
   //Update XCUT status
   "FB_BPSEthLink_ServerA_V1_00_IDB".IN_rgtStatusXCuts[0].dActualCarriagePos_cmm := "FB_CrossCuts_1_V1_00_IDB".tHMR.dCarriagePosition_cmm;
   "FB_BPSEthLink_ServerA_V1_00_IDB".IN_rgtStatusXCuts[0].dDistanceFromSnaproll_cmm := "FB_CrossCuts_1_V1_00_IDB".tHMR.dDistanceFromSnaproll_cmm;
   "FB_BPSEthLink_ServerA_V1_00_IDB".IN_rgtStatusXCuts[0].dStatus := "FB_CrossCuts_1_V1_00_IDB".tHMR.dStatus;
   "FB_BPSEthLink_ServerA_V1_00_IDB".IN_rgtStatusXCuts[0].dXCutActualStatus := "FB_CrossCuts_1_V1_00_IDB".tHMR.dXCutActualStatus;
   IF "FB_CrossCuts_1_V1_00_IDB".tHMR.dXCutActualStatus = 1 THEN
       "FB_BPSEthLink_ServerA_V1_00_IDB".IN_rgtStatusXCuts[0].dStatus := 7;
   END_IF;

   "FB_BPSEthLink_ServerA_V1_00_IDB".IN_rgtStatusXCuts[1].dActualCarriagePos_cmm := "FB_CrossCuts_2_V1_00_IDB".tHMR.dCarriagePosition_cmm;
   "FB_BPSEthLink_ServerA_V1_00_IDB".IN_rgtStatusXCuts[1].dDistanceFromSnaproll_cmm := "FB_CrossCuts_2_V1_00_IDB".tHMR.dDistanceFromSnaproll_cmm;
   "FB_BPSEthLink_ServerA_V1_00_IDB".IN_rgtStatusXCuts[1].dStatus := "FB_CrossCuts_2_V1_00_IDB".tHMR.dStatus;
   "FB_BPSEthLink_ServerA_V1_00_IDB".IN_rgtStatusXCuts[1].dXCutActualStatus := "FB_CrossCuts_2_V1_00_IDB".tHMR.dXCutActualStatus;

   IF "FB_CrossCuts_2_V1_00_IDB".tHMR.dXCutActualStatus = 1 THEN
       "FB_BPSEthLink_ServerA_V1_00_IDB".IN_rgtStatusXCuts[1].dStatus := 7;
   END_IF;

   //Update YCUT status 
   "FB_BPSEthLink_ServerA_V1_00_IDB".IN_rgtStatusYCuts[0].dBridgeStatus := "FB_YCuts1_V1_00_IDB".OUT_tBridgeStatus.dBridgeStatus;
   "FB_BPSEthLink_ServerA_V1_00_IDB".IN_rgtStatusYCuts[0].dDistanceSnapRoll_cmm := "FB_YCuts1_V1_00_IDB".tHMR.dDistanceFromSnaproll_cmm;
   "FB_BPSEthLink_ServerA_V1_00_IDB".IN_rgtStatusYCuts[0].rgdPosition_cmm := "FB_YCuts1_V1_00_IDB".OUT_tBridgeStatus.rgdPosition_cmm;
   "FB_BPSEthLink_ServerA_V1_00_IDB".IN_rgtStatusYCuts[0].rgxFireON := "FB_YCuts1_V1_00_IDB".OUT_tBridgeStatus.rgxFireON;
   "FB_BPSEthLink_ServerA_V1_00_IDB".IN_rgtStatusYCuts[0].rgxHeadProdOn := "FB_YCuts1_V1_00_IDB".OUT_tBridgeStatus.rgxHeadProdOn;

   "FB_BPSEthLink_ServerA_V1_00_IDB".IN_rgtStatusYCuts[1].dBridgeStatus := "FB_YCuts2_V1_00_IDB".OUT_tBridgeStatus.dBridgeStatus;
   "FB_BPSEthLink_ServerA_V1_00_IDB".IN_rgtStatusYCuts[1].dDistanceSnapRoll_cmm := "FB_YCuts2_V1_00_IDB".tHMR.dDistanceFromSnaproll_cmm;
   "FB_BPSEthLink_ServerA_V1_00_IDB".IN_rgtStatusYCuts[1].rgdPosition_cmm := "FB_YCuts2_V1_00_IDB".OUT_tBridgeStatus.rgdPosition_cmm;
   "FB_BPSEthLink_ServerA_V1_00_IDB".IN_rgtStatusYCuts[1].rgxFireON := "FB_YCuts2_V1_00_IDB".OUT_tBridgeStatus.rgxFireON;
   "FB_BPSEthLink_ServerA_V1_00_IDB".IN_rgtStatusYCuts[1].rgxHeadProdOn := "FB_YCuts2_V1_00_IDB".OUT_tBridgeStatus.rgxHeadProdOn;

   //Update general status
   IF (("Z201".ST_xThisPlcActive) AND ("Z201".ST_xPLC1)) THEN
       "FB_BPSEthLink_ServerA_V1_00_IDB".IN_tStatusGeneral.dActivePLC := 1;
   ELSE
       "FB_BPSEthLink_ServerA_V1_00_IDB".IN_tStatusGeneral.dActivePLC := 2;
   END_IF;

   "FB_BPSEthLink_ServerA_V1_00_IDB".IN_tStatusGeneral.dAutoRibSelection := "FB_OptManager_V1_00_IDB".tHMW.dSelectWanderDataSource;
   "FB_BPSEthLink_ServerA_V1_00_IDB".IN_tStatusGeneral.dExtOptSelected := "FB_OptManager_V1_00_IDB".tHMR.dSelOptimizer;
   "FB_BPSEthLink_ServerA_V1_00_IDB".IN_tStatusGeneral.dOptimizerMode := 2;

   IF "FB_OptEthLink_V1_00_IDB".tALM.tS.xCh1NotCon AND "FB_OptEthLink_V1_00_IDB".tALM.tS.xCh2NotCon THEN 
       "FB_BPSEthLink_ServerA_V1_00_IDB".IN_tStatusGeneral.dOptStatus := 1;
   ELSIF "FB_OptEthLink_V1_00_IDB".tALM.tS.xCh1NotCon OR "FB_OptEthLink_V1_00_IDB".tALM.tS.xCh2NotCon THEN
       "FB_BPSEthLink_ServerA_V1_00_IDB".IN_tStatusGeneral.dOptStatus := 7;
   ELSE
       "FB_BPSEthLink_ServerA_V1_00_IDB".IN_tStatusGeneral.dOptStatus := 3;
   END_IF;

   IF "FB_OptManager_V1_00_IDB".tHMW.dSelectWanderDataSource > 0 THEN
       "FB_BPSEthLink_ServerA_V1_00_IDB".IN_tStatusGeneral.dRibbonModality := 1;
   ELSE
       "FB_BPSEthLink_ServerA_V1_00_IDB".IN_tStatusGeneral.dRibbonModality := 4;
   END_IF;

   "FB_BPSEthLink_ServerA_V1_00_IDB".IN_tStatusGeneral.dScanStatus := "FB_ISRA5D_IDB".tHMR.dInspectionStatus;

   IF "FB_OptManager_V1_00_IDB".tHMW.dSelectWanderMode = 0 THEN
       "FB_BPSEthLink_ServerA_V1_00_IDB".IN_tStatusGeneral.dTypeWanderSel := 2;
   ELSE
       "FB_BPSEthLink_ServerA_V1_00_IDB".IN_tStatusGeneral.dTypeWanderSel := 1;
   END_IF;

   "FB_BPSEthLink_ServerA_V1_00_IDB".IN_tStatusGeneral.dYC1WandRec_cmm := "FB_YCuts1_V1_00_IDB".AUX_dActualRecoverWander_cmm;
   "FB_BPSEthLink_ServerA_V1_00_IDB".IN_tStatusGeneral.dYC2WandRec_cmm := "FB_YCuts2_V1_00_IDB".AUX_dActualRecoverWander_cmm;
   "FB_BPSEthLink_ServerA_V1_00_IDB".IN_tStatusGeneral.dWanderRecoveryThr_cmm := "FB_OptManager_V1_00_IDB".tHMW.dWanderRecThr_cmm;

   "FB_BPSEthLink_ServerA_V1_00_IDB".IN_tStatusGeneral.dScanGrossWidth_cmm := "FB_ISRA5D_IDB".tHMR.dCurrentGrossWidth_cmm;
   "FB_BPSEthLink_ServerA_V1_00_IDB".IN_tStatusGeneral.dScanNetWidth_cmm := "FB_ISRA5D_IDB".tHMR.dCurrentNetWidth_cmm;
   "FB_BPSEthLink_ServerA_V1_00_IDB".IN_tStatusGeneral.dScanGrossWander_cmm := "FB_ISRA5D_IDB".tHMR.dCurrentGrossWander_cmm;
   "FB_BPSEthLink_ServerA_V1_00_IDB".IN_tStatusGeneral.dScanNetWander_cmm := "FB_ISRA5D_IDB".tHMR.dCurrentNetWander_cmm;

   "FB_BPSEthLink_ServerA_V1_00_IDB".IN_tStatusGeneral.dCameraGrossWidth_cmm := 0;
   "FB_BPSEthLink_ServerA_V1_00_IDB".IN_tStatusGeneral.dCameraNetWidth_cmm := 0;
   "FB_BPSEthLink_ServerA_V1_00_IDB".IN_tStatusGeneral.dCameraGrossWander_cmm := 0;
   "FB_BPSEthLink_ServerA_V1_00_IDB".IN_tStatusGeneral.dCameraNetWander_cmm := 0;



   //BPS Connection B

   "FB_BPSEthLink_ServerB_V1_00_IDB".IN_tRemoteAddress.ADDR[1] := "IPV4_BPS_SERVERB_IP1";
   "FB_BPSEthLink_ServerB_V1_00_IDB".IN_tRemoteAddress.ADDR[2] := "IPV4_BPS_SERVERB_IP2";
   "FB_BPSEthLink_ServerB_V1_00_IDB".IN_tRemoteAddress.ADDR[3] := "IPV4_BPS_SERVERB_IP3";
   "FB_BPSEthLink_ServerB_V1_00_IDB".IN_tRemoteAddress.ADDR[4] := "IPV4_BPS_SERVERB_IP4";

   "FB_BPSEthLink_ServerB_V1_00_IDB".IN_tStatusEncoder.dActualBTC_cmm := "DB_Encoder".dActualEncoderCounter_cmm;
   "FB_BPSEthLink_ServerB_V1_00_IDB".IN_tStatusEncoder.dTrackSpeed_mm_min := "DB_Encoder".dActSpeedValue_mm_min;

   //Update XCUT status
   "FB_BPSEthLink_ServerB_V1_00_IDB".IN_rgtStatusXCuts[0].dActualCarriagePos_cmm := "FB_CrossCuts_1_V1_00_IDB".tHMR.dCarriagePosition_cmm;
   "FB_BPSEthLink_ServerB_V1_00_IDB".IN_rgtStatusXCuts[0].dDistanceFromSnaproll_cmm := "FB_CrossCuts_1_V1_00_IDB".tHMR.dDistanceFromSnaproll_cmm;
   "FB_BPSEthLink_ServerB_V1_00_IDB".IN_rgtStatusXCuts[0].dStatus := "FB_CrossCuts_1_V1_00_IDB".tHMR.dStatus;
   "FB_BPSEthLink_ServerB_V1_00_IDB".IN_rgtStatusXCuts[0].dXCutActualStatus := "FB_CrossCuts_1_V1_00_IDB".tHMR.dXCutActualStatus;

   IF "FB_CrossCuts_1_V1_00_IDB".tHMR.dXCutActualStatus = 1 THEN
       "FB_BPSEthLink_ServerB_V1_00_IDB".IN_rgtStatusXCuts[0].dStatus := 7;
   END_IF;

   "FB_BPSEthLink_ServerB_V1_00_IDB".IN_rgtStatusXCuts[1].dActualCarriagePos_cmm := "FB_CrossCuts_2_V1_00_IDB".tHMR.dCarriagePosition_cmm;
   "FB_BPSEthLink_ServerB_V1_00_IDB".IN_rgtStatusXCuts[1].dDistanceFromSnaproll_cmm := "FB_CrossCuts_2_V1_00_IDB".tHMR.dDistanceFromSnaproll_cmm;
   "FB_BPSEthLink_ServerB_V1_00_IDB".IN_rgtStatusXCuts[1].dStatus := "FB_CrossCuts_2_V1_00_IDB".tHMR.dStatus;
   "FB_BPSEthLink_ServerB_V1_00_IDB".IN_rgtStatusXCuts[1].dXCutActualStatus := "FB_CrossCuts_2_V1_00_IDB".tHMR.dXCutActualStatus;

   IF "FB_CrossCuts_2_V1_00_IDB".tHMR.dXCutActualStatus = 1 THEN
       "FB_BPSEthLink_ServerB_V1_00_IDB".IN_rgtStatusXCuts[1].dStatus := 7;
   END_IF;

   //Update YCUT status 
   "FB_BPSEthLink_ServerB_V1_00_IDB".IN_rgtStatusYCuts[0].dBridgeStatus := "FB_YCuts1_V1_00_IDB".OUT_tBridgeStatus.dBridgeStatus;
   "FB_BPSEthLink_ServerB_V1_00_IDB".IN_rgtStatusYCuts[0].dDistanceSnapRoll_cmm := "FB_YCuts1_V1_00_IDB".tHMR.dDistanceFromSnaproll_cmm;
   "FB_BPSEthLink_ServerB_V1_00_IDB".IN_rgtStatusYCuts[0].rgdPosition_cmm := "FB_YCuts1_V1_00_IDB".OUT_tBridgeStatus.rgdPosition_cmm;
   "FB_BPSEthLink_ServerB_V1_00_IDB".IN_rgtStatusYCuts[0].rgxFireON := "FB_YCuts1_V1_00_IDB".OUT_tBridgeStatus.rgxFireON;
   "FB_BPSEthLink_ServerB_V1_00_IDB".IN_rgtStatusYCuts[0].rgxHeadProdOn := "FB_YCuts1_V1_00_IDB".OUT_tBridgeStatus.rgxHeadProdOn;

   "FB_BPSEthLink_ServerB_V1_00_IDB".IN_rgtStatusYCuts[1].dBridgeStatus := "FB_YCuts2_V1_00_IDB".OUT_tBridgeStatus.dBridgeStatus;
   "FB_BPSEthLink_ServerB_V1_00_IDB".IN_rgtStatusYCuts[1].dDistanceSnapRoll_cmm := "FB_YCuts2_V1_00_IDB".tHMR.dDistanceFromSnaproll_cmm;
   "FB_BPSEthLink_ServerB_V1_00_IDB".IN_rgtStatusYCuts[1].rgdPosition_cmm := "FB_YCuts2_V1_00_IDB".OUT_tBridgeStatus.rgdPosition_cmm;
   "FB_BPSEthLink_ServerB_V1_00_IDB".IN_rgtStatusYCuts[1].rgxFireON := "FB_YCuts2_V1_00_IDB".OUT_tBridgeStatus.rgxFireON;
   "FB_BPSEthLink_ServerB_V1_00_IDB".IN_rgtStatusYCuts[1].rgxHeadProdOn := "FB_YCuts2_V1_00_IDB".OUT_tBridgeStatus.rgxHeadProdOn;

   //Update general status
   IF (("Z201".ST_xThisPlcActive) AND ("Z201".ST_xPLC1)) THEN
       "FB_BPSEthLink_ServerB_V1_00_IDB".IN_tStatusGeneral.dActivePLC := 1;
   ELSE
       "FB_BPSEthLink_ServerB_V1_00_IDB".IN_tStatusGeneral.dActivePLC := 2;
   END_IF;

   "FB_BPSEthLink_ServerB_V1_00_IDB".IN_tStatusGeneral.dAutoRibSelection := "FB_OptManager_V1_00_IDB".tHMW.dSelectWanderDataSource;
   "FB_BPSEthLink_ServerB_V1_00_IDB".IN_tStatusGeneral.dExtOptSelected := "FB_OptManager_V1_00_IDB".tHMR.dSelOptimizer;
   "FB_BPSEthLink_ServerB_V1_00_IDB".IN_tStatusGeneral.dOptimizerMode := 2;

   IF "FB_OptEthLink_V1_00_IDB".tALM.tS.xCh1NotCon AND "FB_OptEthLink_V1_00_IDB".tALM.tS.xCh2NotCon THEN 
       "FB_BPSEthLink_ServerB_V1_00_IDB".IN_tStatusGeneral.dOptStatus := 1;
   ELSIF "FB_OptEthLink_V1_00_IDB".tALM.tS.xCh1NotCon OR "FB_OptEthLink_V1_00_IDB".tALM.tS.xCh2NotCon THEN
       "FB_BPSEthLink_ServerB_V1_00_IDB".IN_tStatusGeneral.dOptStatus := 7;
   ELSE
       "FB_BPSEthLink_ServerB_V1_00_IDB".IN_tStatusGeneral.dOptStatus := 3;
   END_IF;

   IF "FB_OptManager_V1_00_IDB".tHMW.dSelectWanderDataSource > 0 THEN
       "FB_BPSEthLink_ServerB_V1_00_IDB".IN_tStatusGeneral.dRibbonModality := 1;
   ELSE
       "FB_BPSEthLink_ServerB_V1_00_IDB".IN_tStatusGeneral.dRibbonModality := 4;
   END_IF;

   "FB_BPSEthLink_ServerB_V1_00_IDB".IN_tStatusGeneral.dScanStatus := "FB_ISRA5D_IDB".tHMR.dInspectionStatus;

   IF "FB_OptManager_V1_00_IDB".tHMW.dSelectWanderMode = 0 THEN
       "FB_BPSEthLink_ServerB_V1_00_IDB".IN_tStatusGeneral.dTypeWanderSel := 2;
   ELSE
       "FB_BPSEthLink_ServerB_V1_00_IDB".IN_tStatusGeneral.dTypeWanderSel := 1;
   END_IF;

   "FB_BPSEthLink_ServerB_V1_00_IDB".IN_tStatusGeneral.dYC1WandRec_cmm := "FB_YCuts1_V1_00_IDB".AUX_dActualRecoverWander_cmm;
   "FB_BPSEthLink_ServerB_V1_00_IDB".IN_tStatusGeneral.dYC2WandRec_cmm := "FB_YCuts2_V1_00_IDB".AUX_dActualRecoverWander_cmm;
   "FB_BPSEthLink_ServerB_V1_00_IDB".IN_tStatusGeneral.dWanderRecoveryThr_cmm := "FB_OptManager_V1_00_IDB".tHMW.dWanderRecThr_cmm;

   "FB_BPSEthLink_ServerB_V1_00_IDB".IN_tStatusGeneral.dScanGrossWidth_cmm := "FB_ISRA5D_IDB".tHMR.dCurrentGrossWidth_cmm;
   "FB_BPSEthLink_ServerB_V1_00_IDB".IN_tStatusGeneral.dScanNetWidth_cmm := "FB_ISRA5D_IDB".tHMR.dCurrentNetWidth_cmm;
   "FB_BPSEthLink_ServerB_V1_00_IDB".IN_tStatusGeneral.dScanGrossWander_cmm := "FB_ISRA5D_IDB".tHMR.dCurrentGrossWander_cmm;
   "FB_BPSEthLink_ServerB_V1_00_IDB".IN_tStatusGeneral.dScanNetWander_cmm := "FB_ISRA5D_IDB".tHMR.dCurrentNetWander_cmm;

   "FB_BPSEthLink_ServerB_V1_00_IDB".IN_tStatusGeneral.dCameraGrossWidth_cmm := 0;
   "FB_BPSEthLink_ServerB_V1_00_IDB".IN_tStatusGeneral.dCameraNetWidth_cmm := 0;
   "FB_BPSEthLink_ServerB_V1_00_IDB".IN_tStatusGeneral.dCameraGrossWander_cmm := 0;
   "FB_BPSEthLink_ServerB_V1_00_IDB".IN_tStatusGeneral.dCameraNetWander_cmm := 0;
END_REGION

REGION Network 4: BPS A Connection data
   RUNG wire#powerrail
      "FB_BPSEthLink_ServerA_V1_00_IDB"(IN_xBPSServerA := TRUE, IN_xCycleON :=, IN_xCycleONDel := "Z201".ST_xCycleONDelayed, IN_xGeneralReset := "Z201".ST_xMachineReset, IN_xResetAlarms := "Z201".tmOFF_ResetAlarm.OUT_xDone, IN_xFaultsEnabled := "Z201".ST_xFaultsEnabled, IN_xThisPLCActive := "Z201".ST_xThisPlcActive, IN_dLineSpeed_mm_min := "FB_CommunicationZ300_V1.00_DB".IN_tIDeviceDataIN.Z300.dLineSpeed_mm_min, IN_tStatusGeneral :=, IN_tStatusEncoder :=, IN_tStatusDigitizer_1 :=, IN_tStatusDigitizer_2 :=, IN_rgtStatusXCuts :=, IN_rgtStatusYCuts :=, IN_rgtStatusMarkers :=, IN_tInterfaceID := "Local~PROFINET_MCC1200", IN_tID := "CONNUOC_BPS_SERVERA", IN_tRemoteAddress :=, IN_uiRemotePort := "UINT_BPS_SERVERA_PORT", INO_tCaps := "DB_Plates", INO_tInitialize := "GP_OB_Initialize_Main_IDB", INO_tDefects := "DB_Defects".THIS, INO_tMessages := "RP_Message".tTankMessageForReport, INO_tAddMessageFromOpt := "RP_Message".MexFromOptimizer.tAddMessageFromOptTaskMain, INO_tRibbon := "DB_RibbonData", INO_xMessageAnomaly := "RP_Message".tALM.tS.xMessageAnomaly)
   END_RUNG
   // the same network as SCL:
   "FB_BPSEthLink_ServerA_V1_00_IDB"(IN_xBPSServerA := TRUE,   // "FB_BPSEthLink_V1.00"
                           IN_xCycleONDel := "Z201".ST_xCycleONDelayed,
                           IN_xGeneralReset := "Z201".ST_xMachineReset,
                           IN_xResetAlarms := "Z201".tmOFF_ResetAlarm.OUT_xDone,
                           IN_xFaultsEnabled := "Z201".ST_xFaultsEnabled,
                           IN_xThisPLCActive := "Z201".ST_xThisPlcActive,
                           IN_dLineSpeed_mm_min := "FB_CommunicationZ300_V1.00_DB".IN_tIDeviceDataIN.Z300.dLineSpeed_mm_min,
                           IN_tInterfaceID := "Local~PROFINET_MCC1200",
                           IN_tID := "CONNUOC_BPS_SERVERA",
                           IN_uiRemotePort := "UINT_BPS_SERVERA_PORT",
                           INO_tCaps := "DB_Plates",
                           INO_tInitialize := "GP_OB_Initialize_Main_IDB",
                           INO_tDefects := "DB_Defects".THIS,
                           INO_tMessages := "RP_Message".tTankMessageForReport,
                           INO_tAddMessageFromOpt := "RP_Message".MexFromOptimizer.tAddMessageFromOptTaskMain,
                           INO_tRibbon := "DB_RibbonData",
                           INO_xMessageAnomaly := "RP_Message".tALM.tS.xMessageAnomaly);
END_REGION

REGION Network 5: BPS B Connection data
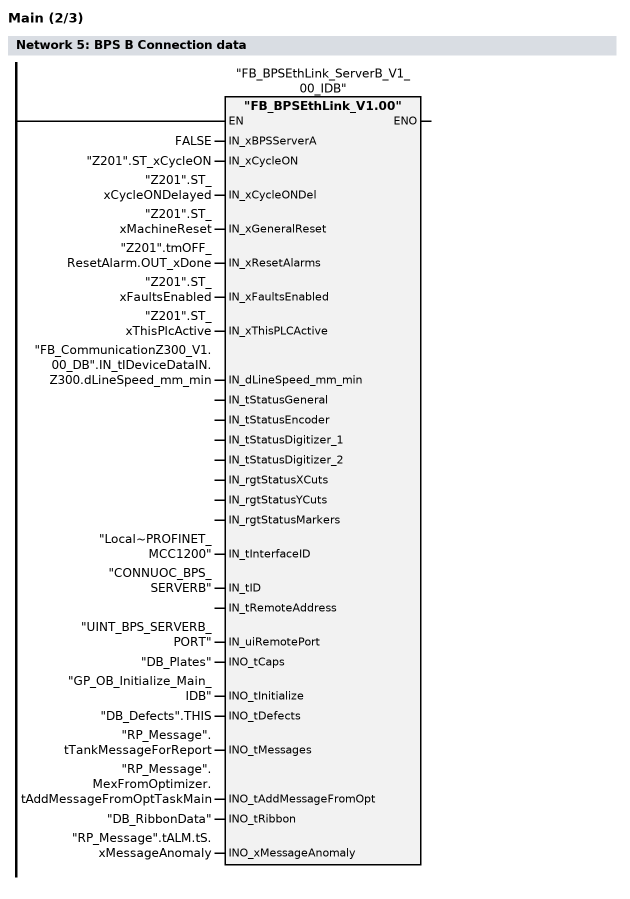
   RUNG wire#powerrail
      "FB_BPSEthLink_ServerB_V1_00_IDB"(IN_xBPSServerA := FALSE, IN_xCycleON := "Z201".ST_xCycleON, IN_xCycleONDel := "Z201".ST_xCycleONDelayed, IN_xGeneralReset := "Z201".ST_xMachineReset, IN_xResetAlarms := "Z201".tmOFF_ResetAlarm.OUT_xDone, IN_xFaultsEnabled := "Z201".ST_xFaultsEnabled, IN_xThisPLCActive := "Z201".ST_xThisPlcActive, IN_dLineSpeed_mm_min := "FB_CommunicationZ300_V1.00_DB".IN_tIDeviceDataIN.Z300.dLineSpeed_mm_min, IN_tStatusGeneral :=, IN_tStatusEncoder :=, IN_tStatusDigitizer_1 :=, IN_tStatusDigitizer_2 :=, IN_rgtStatusXCuts :=, IN_rgtStatusYCuts :=, IN_rgtStatusMarkers :=, IN_tInterfaceID := "Local~PROFINET_MCC1200", IN_tID := "CONNUOC_BPS_SERVERB", IN_tRemoteAddress :=, IN_uiRemotePort := "UINT_BPS_SERVERB_PORT", INO_tCaps := "DB_Plates", INO_tInitialize := "GP_OB_Initialize_Main_IDB", INO_tDefects := "DB_Defects".THIS, INO_tMessages := "RP_Message".tTankMessageForReport, INO_tAddMessageFromOpt := "RP_Message".MexFromOptimizer.tAddMessageFromOptTaskMain, INO_tRibbon := "DB_RibbonData", INO_xMessageAnomaly := "RP_Message".tALM.tS.xMessageAnomaly)
   END_RUNG
   // the same network as SCL:
   "FB_BPSEthLink_ServerB_V1_00_IDB"(IN_xBPSServerA := FALSE,   // "FB_BPSEthLink_V1.00"
                           IN_xCycleON := "Z201".ST_xCycleON,
                           IN_xCycleONDel := "Z201".ST_xCycleONDelayed,
                           IN_xGeneralReset := "Z201".ST_xMachineReset,
                           IN_xResetAlarms := "Z201".tmOFF_ResetAlarm.OUT_xDone,
                           IN_xFaultsEnabled := "Z201".ST_xFaultsEnabled,
                           IN_xThisPLCActive := "Z201".ST_xThisPlcActive,
                           IN_dLineSpeed_mm_min := "FB_CommunicationZ300_V1.00_DB".IN_tIDeviceDataIN.Z300.dLineSpeed_mm_min,
                           IN_tInterfaceID := "Local~PROFINET_MCC1200",
                           IN_tID := "CONNUOC_BPS_SERVERB",
                           IN_uiRemotePort := "UINT_BPS_SERVERB_PORT",
                           INO_tCaps := "DB_Plates",
                           INO_tInitialize := "GP_OB_Initialize_Main_IDB",
                           INO_tDefects := "DB_Defects".THIS,
                           INO_tMessages := "RP_Message".tTankMessageForReport,
                           INO_tAddMessageFromOpt := "RP_Message".MexFromOptimizer.tAddMessageFromOptTaskMain,
                           INO_tRibbon := "DB_RibbonData",
                           INO_xMessageAnomaly := "RP_Message".tALM.tS.xMessageAnomaly);
END_REGION

REGION Network 6 (SCL): Optimizer connection data
   //Update YCUT status 
   "FB_OptEthLink_V1_00_IDB".IN_rgtStatusYCuts[0].dBridgeStatus := "FB_YCuts1_V1_00_IDB".OUT_tBridgeStatus.dBridgeStatus;
   "FB_OptEthLink_V1_00_IDB".IN_rgtStatusYCuts[0].dDistanceSnapRoll_cmm := "FB_YCuts1_V1_00_IDB".tHMR.dDistanceFromSnaproll_cmm;
   "FB_OptEthLink_V1_00_IDB".IN_rgtStatusYCuts[0].rgdPosition_cmm := "FB_YCuts1_V1_00_IDB".OUT_tBridgeStatus.rgdPosition_cmm;
   "FB_OptEthLink_V1_00_IDB".IN_rgtStatusYCuts[0].rgxFireON := "FB_YCuts1_V1_00_IDB".OUT_tBridgeStatus.rgxFireON;
   "FB_OptEthLink_V1_00_IDB".IN_rgtStatusYCuts[0].rgxHeadProdOn := "FB_YCuts1_V1_00_IDB".OUT_tBridgeStatus.rgxHeadProdOn;


   "FB_OptEthLink_V1_00_IDB".IN_rgtStatusYCuts[1].dBridgeStatus := "FB_YCuts2_V1_00_IDB".OUT_tBridgeStatus.dBridgeStatus;
   "FB_OptEthLink_V1_00_IDB".IN_rgtStatusYCuts[1].dDistanceSnapRoll_cmm := "FB_YCuts2_V1_00_IDB".tHMR.dDistanceFromSnaproll_cmm;
   "FB_OptEthLink_V1_00_IDB".IN_rgtStatusYCuts[1].rgdPosition_cmm := "FB_YCuts2_V1_00_IDB".OUT_tBridgeStatus.rgdPosition_cmm;
   "FB_OptEthLink_V1_00_IDB".IN_rgtStatusYCuts[1].rgxFireON := "FB_YCuts2_V1_00_IDB".OUT_tBridgeStatus.rgxFireON;
   "FB_OptEthLink_V1_00_IDB".IN_rgtStatusYCuts[1].rgxHeadProdOn := "FB_YCuts2_V1_00_IDB".OUT_tBridgeStatus.rgxHeadProdOn;
   "FB_OptEthLink_V1_00_IDB".IN_rgtStatusXCuts[0].dActualCarriagePos_cmm := "FB_CrossCuts_1_V1_00_IDB".tHMR.dCarriagePosition_cmm;
   "FB_OptEthLink_V1_00_IDB".IN_rgtStatusXCuts[0].dDistanceFromSnaproll_cmm := "FB_CrossCuts_1_V1_00_IDB".tHMR.dDistanceFromSnaproll_cmm;
   "FB_OptEthLink_V1_00_IDB".IN_rgtStatusXCuts[0].dStatus := "FB_CrossCuts_1_V1_00_IDB".tHMR.dStatus;
   "FB_OptEthLink_V1_00_IDB".IN_rgtStatusXCuts[0].dXCutActualStatus := "FB_CrossCuts_1_V1_00_IDB".tHMR.dXCutActualStatus;
   "FB_OptEthLink_V1_00_IDB".IN_rgtStatusXCuts[0].dCutTime_ms := "FB_CrossCuts_1_V1_00_IDB".AUX_dCutTime100Per_ms;

   "FB_OptEthLink_V1_00_IDB".IN_rgtStatusXCuts[1].dActualCarriagePos_cmm := "FB_CrossCuts_2_V1_00_IDB".tHMR.dCarriagePosition_cmm;
   "FB_OptEthLink_V1_00_IDB".IN_rgtStatusXCuts[1].dDistanceFromSnaproll_cmm := "FB_CrossCuts_2_V1_00_IDB".tHMR.dDistanceFromSnaproll_cmm;
   "FB_OptEthLink_V1_00_IDB".IN_rgtStatusXCuts[1].dStatus := "FB_CrossCuts_2_V1_00_IDB".tHMR.dStatus;
   "FB_OptEthLink_V1_00_IDB".IN_rgtStatusXCuts[1].dXCutActualStatus := "FB_CrossCuts_2_V1_00_IDB".tHMR.dXCutActualStatus;
   "FB_OptEthLink_V1_00_IDB".IN_rgtStatusXCuts[1].dCutTime_ms := "FB_CrossCuts_2_V1_00_IDB".AUX_dCutTime100Per_ms;

   "FB_OptEthLink_V1_00_IDB".IN_rgtStatusXCuts[2].dActualCarriagePos_cmm := 0;
   "FB_OptEthLink_V1_00_IDB".IN_rgtStatusXCuts[2].dDistanceFromSnaproll_cmm := 0;
   "FB_OptEthLink_V1_00_IDB".IN_rgtStatusXCuts[2].dStatus := 1;
   "FB_OptEthLink_V1_00_IDB".IN_rgtStatusXCuts[2].dXCutActualStatus := 1;
   "FB_OptEthLink_V1_00_IDB".IN_rgtStatusXCuts[2].dCutTime_ms := 0;

   "FB_OptEthLink_V1_00_IDB".IN_rgtStatusXCuts[3].dActualCarriagePos_cmm := 0;
   "FB_OptEthLink_V1_00_IDB".IN_rgtStatusXCuts[3].dDistanceFromSnaproll_cmm := 0;
   "FB_OptEthLink_V1_00_IDB".IN_rgtStatusXCuts[3].dStatus :=1;
   "FB_OptEthLink_V1_00_IDB".IN_rgtStatusXCuts[3].dXCutActualStatus := 1;
   "FB_OptEthLink_V1_00_IDB".IN_rgtStatusXCuts[3].dCutTime_ms := 0;

   "FB_OptEthLink_V1_00_IDB".IN_rgtStatusMarker[3].dBridgeProdModeActual := 0;
   "FB_OptEthLink_V1_00_IDB".IN_rgtStatusMarker[3].dDistanceFromCenterLine_cmm := 0;
   "FB_OptEthLink_V1_00_IDB".IN_rgtStatusMarker[3].dDistanceFromSnaproll_cmm := 0;
   "FB_OptEthLink_V1_00_IDB".IN_rgtStatusMarker[3].dHeadPosition_cmm := 0;
   "FB_OptEthLink_V1_00_IDB".IN_rgtStatusMarker[3].dSpraySpace_cmm := 0;

   "FB_OptEthLink_V1_00_IDB".IN_rgtStatusMarker[4].dBridgeProdModeActual := 0;
   "FB_OptEthLink_V1_00_IDB".IN_rgtStatusMarker[4].dDistanceFromCenterLine_cmm := 0;
   "FB_OptEthLink_V1_00_IDB".IN_rgtStatusMarker[4].dDistanceFromSnaproll_cmm := 0;
   "FB_OptEthLink_V1_00_IDB".IN_rgtStatusMarker[4].dHeadPosition_cmm := 0;
   "FB_OptEthLink_V1_00_IDB".IN_rgtStatusMarker[4].dSpraySpace_cmm := 0;
END_REGION

REGION Network 7: Optimizer connection
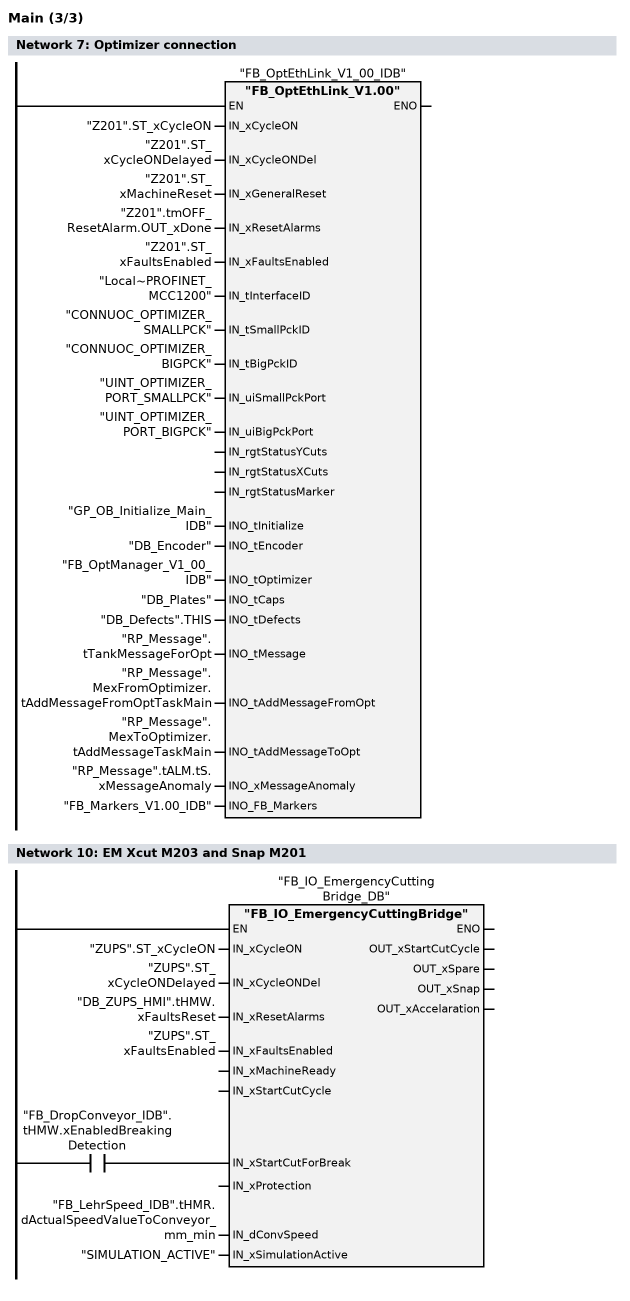
   RUNG wire#powerrail
      "FB_OptEthLink_V1_00_IDB"(IN_xCycleON := "Z201".ST_xCycleON, IN_xCycleONDel := "Z201".ST_xCycleONDelayed, IN_xGeneralReset := "Z201".ST_xMachineReset, IN_xResetAlarms := "Z201".tmOFF_ResetAlarm.OUT_xDone, IN_xFaultsEnabled := "Z201".ST_xFaultsEnabled, IN_tInterfaceID := "Local~PROFINET_MCC1200", IN_tSmallPckID := "CONNUOC_OPTIMIZER_SMALLPCK", IN_tBigPckID := "CONNUOC_OPTIMIZER_BIGPCK", IN_uiSmallPckPort := "UINT_OPTIMIZER_PORT_SMALLPCK", IN_uiBigPckPort := "UINT_OPTIMIZER_PORT_BIGPCK", IN_rgtStatusYCuts :=, IN_rgtStatusXCuts :=, IN_rgtStatusMarker :=, INO_tInitialize := "GP_OB_Initialize_Main_IDB", INO_tEncoder := "DB_Encoder", INO_tOptimizer := "FB_OptManager_V1_00_IDB", INO_tCaps := "DB_Plates", INO_tDefects := "DB_Defects".THIS, INO_tMessage := "RP_Message".tTankMessageForOpt, INO_tAddMessageFromOpt := "RP_Message".MexFromOptimizer.tAddMessageFromOptTaskMain, INO_tAddMessageToOpt := "RP_Message".MexToOptimizer.tAddMessageTaskMain, INO_xMessageAnomaly := "RP_Message".tALM.tS.xMessageAnomaly, INO_FB_Markers := "FB_Markers_V1.00_IDB")
   END_RUNG
   // the same network as SCL:
   "FB_OptEthLink_V1_00_IDB"(IN_xCycleON := "Z201".ST_xCycleON,   // "FB_OptEthLink_V1.00"
                           IN_xCycleONDel := "Z201".ST_xCycleONDelayed,
                           IN_xGeneralReset := "Z201".ST_xMachineReset,
                           IN_xResetAlarms := "Z201".tmOFF_ResetAlarm.OUT_xDone,
                           IN_xFaultsEnabled := "Z201".ST_xFaultsEnabled,
                           IN_tInterfaceID := "Local~PROFINET_MCC1200",
                           IN_tSmallPckID := "CONNUOC_OPTIMIZER_SMALLPCK",
                           IN_tBigPckID := "CONNUOC_OPTIMIZER_BIGPCK",
                           IN_uiSmallPckPort := "UINT_OPTIMIZER_PORT_SMALLPCK",
                           IN_uiBigPckPort := "UINT_OPTIMIZER_PORT_BIGPCK",
                           INO_tInitialize := "GP_OB_Initialize_Main_IDB",
                           INO_tEncoder := "DB_Encoder",
                           INO_tOptimizer := "FB_OptManager_V1_00_IDB",
                           INO_tCaps := "DB_Plates",
                           INO_tDefects := "DB_Defects".THIS,
                           INO_tMessage := "RP_Message".tTankMessageForOpt,
                           INO_tAddMessageFromOpt := "RP_Message".MexFromOptimizer.tAddMessageFromOptTaskMain,
                           INO_tAddMessageToOpt := "RP_Message".MexToOptimizer.tAddMessageTaskMain,
                           INO_xMessageAnomaly := "RP_Message".tALM.tS.xMessageAnomaly,
                           INO_FB_Markers := "FB_Markers_V1.00_IDB");
END_REGION

REGION Network 8: FRom Z201
END_REGION

REGION Network 9 (SCL)

   "InputZ201_Idevice"();

   "ZUPS_Faults"();
   "ZUPS_Logics"();
   "ZUPS_Output"();

   "Z201_Faults"();
   "Z201_Logics"();
   "Z201_Output"();

   "SCADA_Mapping"();





   "FB_DropConveyor_IDB"(IN_xCycleON := "Z201".ST_xCycleON  AND "ZUPS".ST_xCycleON,
                         IN_xCycleONDel := "Z201".ST_xCycleONDelayed,
                         IN_xResetAlarms := "ZUPS".tmOFF_ResetAlarm.OUT_xDone,
                         IN_xFaultsEnabled := "ZUPS".ST_xFaultsEnabled,
                         IN_xManualMode := "FB_Z200Conveyor_M204_IDB".tHMR.xManualCommandEnabled,
                         IN_dActualLehrSpeed_mm_min :="FB_LehrSpeed_IDB".tHMR.dActualSpeedValueToConveyor_mm_min,
                         IN_dGlassBreakMachineIndex := "DGLASSBREAKMACHINEINDEX_M204",
                         IN_dGlassBreakGetIndex := "DGLASSBREAKGET_M204",
                         IN_xSimulationActive := "SIMULATION_ACTIVE",
                         INO_tRibbon := "DB_RibbonData");

   "FB_BreakerM206_V1_00_IDB"(IN_xCycleON := "ZUPS".ST_xCycleON,
                              IN_xCycleONDel := "ZUPS".ST_xCycleONDelayed,
                              IN_xGeneralReset := "Z201".ST_xMachineReset,
                              IN_xResetAlarms := "ZUPS".tmOFF_ResetAlarm.OUT_xDone,
                              IN_xFaultsEnabled := "ZUPS".ST_xFaultsEnabled,
                              IN_xDropConveyorDown := "FB_DropConveyor_IDB".tHMR.xDownPosition,
                              INO_tOBInitialize := "GP_OB_Initialize_Main_IDB");
END_REGION

REGION Network 10: EM Xcut M203 and Snap M201
   RUNG wire#powerrail
      "FB_IO_EmergencyCuttingBridge_DB"(IN_xStartCutForBreak := wire#w1, IN_xCycleON := "ZUPS".ST_xCycleON, IN_xCycleONDel := "ZUPS".ST_xCycleONDelayed, IN_xResetAlarms := "DB_ZUPS_HMI".tHMW.xFaultsReset, IN_xFaultsEnabled := "ZUPS".ST_xFaultsEnabled, IN_xMachineReady :=, IN_xStartCutCycle :=, IN_xProtection :=, IN_dConvSpeed := "FB_LehrSpeed_IDB".tHMR.dActualSpeedValueToConveyor_mm_min, IN_xSimulationActive := "SIMULATION_ACTIVE", OUT_xStartCutCycle =>, OUT_xSpare =>, OUT_xSnap =>, OUT_xAccelaration =>)
   END_RUNG
   RUNG wire#powerrail
      Contact( "FB_DropConveyor_IDB".tHMW.xEnabledBreakingDetection )
   END_RUNG wire#w1
   // the same network as SCL:
   "FB_IO_EmergencyCuttingBridge_DB"(IN_xCycleON := "ZUPS".ST_xCycleON,   // "FB_IO_EmergencyCuttingBridge"
                           IN_xCycleONDel := "ZUPS".ST_xCycleONDelayed,
                           IN_xResetAlarms := "DB_ZUPS_HMI".tHMW.xFaultsReset,
                           IN_xFaultsEnabled := "ZUPS".ST_xFaultsEnabled,
                           IN_xStartCutForBreak := "FB_DropConveyor_IDB".tHMW.xEnabledBreakingDetection,
                           IN_dConvSpeed := "FB_LehrSpeed_IDB".tHMR.dActualSpeedValueToConveyor_mm_min,
                           IN_xSimulationActive := "SIMULATION_ACTIVE");
END_REGION

REGION Network 11 (SCL): Z200 Conveyors
   "Z200SinamicsCU_Management"();

   //M201
   //motor Config 
   #TMP_rgtMotorConfig.iIOAddress_MM := 2020;
   #TMP_rgtMotorConfig.iPZD_MM := 1;
   #TMP_rgtMotorConfig.dMaxSpeed_rpm := 3000;
   #TMP_rgtMotorConfig.rK_rpm_mmMin := 15.7080;
   #TMP_rgtMotorConfig.rK_mmMin_Rpm := 0.063661977;
   #TMP_rgtMotorConfig.rMaxAcc := 3.142;
   #TMP_rgtMotorConfig.rMaxDec := 3.142;
   #TMP_rgtMotorConfig.rAcc := 3.142;
   #TMP_rgtMotorConfig.rDec := 3.142;
   #TMP_rgtMotorConfig.xModuleCorrect := TRUE;
   #TMP_rgtMotorConfig.xMDI_Continue := TRUE;



   "FB_Z200Conveyor_M201_IDB"(IN_xCycleON := "ZUPS".ST_xCycleON,
                              IN_xCycleONDel := "ZUPS".ST_xCycleONDelayed,
                              IN_xFaultsEnabled := "ZUPS".ST_xFaultsEnabled,
                              IN_xResetAlarms := "Z201".tmOFF_ResetAlarm.OUT_xDone,
                              IN_xAccelation:=FALSE,
                              IN_rgtMotorConfig := #TMP_rgtMotorConfig);

   //M204
   //motor Config 
   #TMP_rgtMotorConfig.iIOAddress_MM := 2050;
   #TMP_rgtMotorConfig.iPZD_MM := 1;
   #TMP_rgtMotorConfig.dMaxSpeed_rpm := 3000;
   #TMP_rgtMotorConfig.rK_rpm_mmMin := 15.7080;
   #TMP_rgtMotorConfig.rK_mmMin_Rpm := 0.063661977;
   #TMP_rgtMotorConfig.rMaxAcc := 3.142;
   #TMP_rgtMotorConfig.rMaxDec := 3.142;
   #TMP_rgtMotorConfig.rAcc := 3.142;
   #TMP_rgtMotorConfig.rDec := 3.142;
   #TMP_rgtMotorConfig.xModuleCorrect := TRUE;
   #TMP_rgtMotorConfig.xMDI_Continue := TRUE;

   "FB_Z200Conveyor_M204_IDB"(IN_xCycleON:="ZUPS".ST_xCycleON,
                              IN_xCycleONDel:="ZUPS".ST_xCycleONDelayed,
                              IN_xResetAlarms:="ZUPS".ST_xFaultsEnabled,
                              IN_xFaultsEnabled:= "Z201".tmOFF_ResetAlarm.OUT_xDone,
                              IN_xAccelation:="FB_IO_EmergencyCuttingBridge_DB".OUT_xAccelaration AND "FB_DropConveyor_IDB".INPUT.xDownPosition ,
                              IN_rgtMotorConfig:= #TMP_rgtMotorConfig);



   //M205
   //motor Config 
   #TMP_rgtMotorConfig.iIOAddress_MM := 2080;
   #TMP_rgtMotorConfig.iPZD_MM := 1;
   #TMP_rgtMotorConfig.dMaxSpeed_rpm := 3000;
   #TMP_rgtMotorConfig.rK_rpm_mmMin := 50.05650478;
   #TMP_rgtMotorConfig.rK_mmMin_Rpm := 0.019977424;
   #TMP_rgtMotorConfig.rMaxAcc := 3.575;
   #TMP_rgtMotorConfig.rMaxDec :=  3.575;
   #TMP_rgtMotorConfig.rAcc :=  3.575;
   #TMP_rgtMotorConfig.rDec :=  3.575;
   #TMP_rgtMotorConfig.xModuleCorrect := TRUE;
   #TMP_rgtMotorConfig.xMDI_Continue := TRUE;



   "FB_Z200Conveyor_M205_IDB"(IN_xCycleON := "ZUPS".ST_xCycleON,
                              IN_xCycleONDel := "ZUPS".ST_xCycleONDelayed,
                              IN_xFaultsEnabled := "ZUPS".ST_xFaultsEnabled,
                              IN_xResetAlarms := "Z201".tmOFF_ResetAlarm.OUT_xDone,
                              IN_xAccelation:=FALSE,
                              IN_rgtMotorConfig := #TMP_rgtMotorConfig);

   //M214
   //motor Config 
   #TMP_rgtMotorConfig.iIOAddress_MM := 2220;
   #TMP_rgtMotorConfig.iPZD_MM := 1;
   #TMP_rgtMotorConfig.dMaxSpeed_rpm := 3000;
   #TMP_rgtMotorConfig.rK_rpm_mmMin := 15.7080;
   #TMP_rgtMotorConfig.rK_mmMin_Rpm := 0.063661977;
   #TMP_rgtMotorConfig.rMaxAcc := 3.142;
   #TMP_rgtMotorConfig.rMaxDec := 3.142;
   #TMP_rgtMotorConfig.rAcc := 3.142;
   #TMP_rgtMotorConfig.rDec := 3.142;
   #TMP_rgtMotorConfig.xModuleCorrect := TRUE;
   #TMP_rgtMotorConfig.xMDI_Continue := TRUE;


   "FB_Z200Conveyor_M214_iDB"(IN_xCycleON := "Z201".ST_xCycleON,
                              IN_xCycleONDel := "Z201".ST_xCycleONDelayed,
                              IN_xFaultsEnabled := "Z201".ST_xFaultsEnabled,
                              IN_xResetAlarms := "Z201".tmOFF_ResetAlarm.OUT_xDone,
                              IN_xAccelation:=FALSE,
                              IN_rgtMotorConfig := #TMP_rgtMotorConfig);

   //M218
   //motor Config 
   #TMP_rgtMotorConfig.iIOAddress_MM := 2270;
   #TMP_rgtMotorConfig.iPZD_MM := 1;
   #TMP_rgtMotorConfig.dMaxSpeed_rpm := 3000;
   #TMP_rgtMotorConfig.rK_rpm_mmMin := 15.7080;
   #TMP_rgtMotorConfig.rK_mmMin_Rpm := 0.063661977;
   #TMP_rgtMotorConfig.rMaxAcc := 3.142;
   #TMP_rgtMotorConfig.rMaxDec := 3.142;
   #TMP_rgtMotorConfig.rAcc := 3.142;
   #TMP_rgtMotorConfig.rDec := 3.142;
   #TMP_rgtMotorConfig.xModuleCorrect := TRUE;
   #TMP_rgtMotorConfig.xMDI_Continue := TRUE;


   "FB_Z200Conveyor_M218_IDB"(IN_xCycleON := "Z201".ST_xCycleON,
                              IN_xCycleONDel := "Z201".ST_xCycleONDelayed,
                              IN_xFaultsEnabled := "Z201".ST_xFaultsEnabled,
                              IN_xResetAlarms := "Z201".tmOFF_ResetAlarm.OUT_xDone,
                              IN_xAccelation:=FALSE,
                              IN_rgtMotorConfig := #TMP_rgtMotorConfig);



   //M208
   //motor Config 
   #TMP_rgtMotorConfig.iIOAddress_MM := 2320;
   #TMP_rgtMotorConfig.iPZD_MM := 1;
   #TMP_rgtMotorConfig.dMaxSpeed_rpm := 3000;
   #TMP_rgtMotorConfig.rK_rpm_mmMin := 15.7080;
   #TMP_rgtMotorConfig.rK_mmMin_Rpm := 0.063661977;
   #TMP_rgtMotorConfig.rMaxAcc := 3.142;
   #TMP_rgtMotorConfig.rMaxDec := 3.142;
   #TMP_rgtMotorConfig.rAcc := 3.142;
   #TMP_rgtMotorConfig.rDec := 3.142;
   #TMP_rgtMotorConfig.xModuleCorrect := TRUE;
   #TMP_rgtMotorConfig.xMDI_Continue := TRUE;


   "FB_Z200Conveyor_M208_IDB"(IN_xCycleON := "Z201".ST_xCycleON,
                              IN_xCycleONDel := "Z201".ST_xCycleONDelayed,
                              IN_xFaultsEnabled := "Z201".ST_xFaultsEnabled,
                              IN_xResetAlarms := "Z201".tmOFF_ResetAlarm.OUT_xDone,
                              IN_xAccelation:=FALSE,
                              IN_rgtMotorConfig := #TMP_rgtMotorConfig);


   //M211
   //motor Config 
   #TMP_rgtMotorConfig.iIOAddress_MM := 2370;
   #TMP_rgtMotorConfig.iPZD_MM := 1;
   #TMP_rgtMotorConfig.dMaxSpeed_rpm := 3000;
   #TMP_rgtMotorConfig.rK_rpm_mmMin := 15.7080;
   #TMP_rgtMotorConfig.rK_mmMin_Rpm := 0.063661977;
   #TMP_rgtMotorConfig.rMaxAcc := 3.142;
   #TMP_rgtMotorConfig.rMaxDec := 3.142;
   #TMP_rgtMotorConfig.rAcc := 3.142;
   #TMP_rgtMotorConfig.rDec := 3.142;
   #TMP_rgtMotorConfig.xModuleCorrect := TRUE;
   #TMP_rgtMotorConfig.xMDI_Continue := TRUE;



